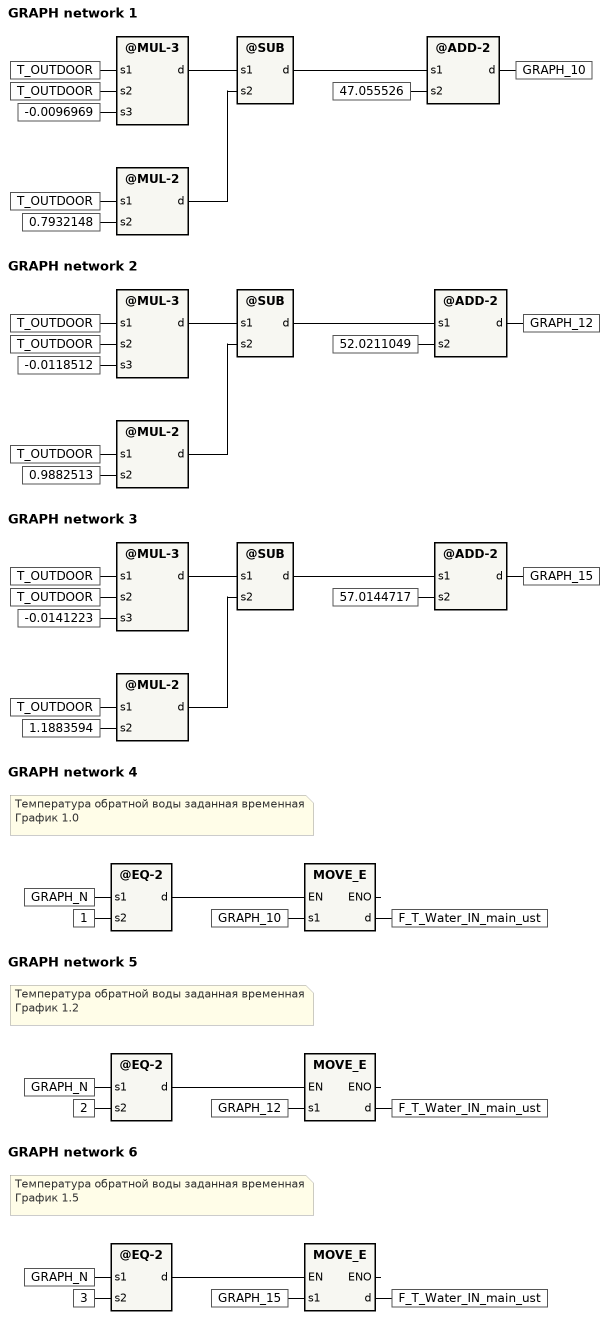
(* network 1 *)
GRAPH_10 := @ADD-2(@SUB(@MUL-3(T_OUTDOOR, T_OUTDOOR, -0.0096969), @MUL-2(T_OUTDOOR, 0.7932148)), 47.055526);
(* network 2 *)
GRAPH_12 := @ADD-2(@SUB(@MUL-3(T_OUTDOOR, T_OUTDOOR, -0.0118512), @MUL-2(T_OUTDOOR, 0.9882513)), 52.0211049);
(* network 3 *)
GRAPH_15 := @ADD-2(@SUB(@MUL-3(T_OUTDOOR, T_OUTDOOR, -0.0141223), @MUL-2(T_OUTDOOR, 1.1883594)), 57.0144717);
(* network 4 *)
(* Температура обратной воды заданная временная График 1.0 *)
MOVE_E(@EQ-2(GRAPH_N, 1), GRAPH_10, F_T_Water_IN_main_ust);
(* network 5 *)
(* Температура обратной воды заданная временная График 1.2 *)
MOVE_E(@EQ-2(GRAPH_N, 2), GRAPH_12, F_T_Water_IN_main_ust);
(* network 6 *)
(* Температура обратной воды заданная временная График 1.5 *)
MOVE_E(@EQ-2(GRAPH_N, 3), GRAPH_15, F_T_Water_IN_main_ust);
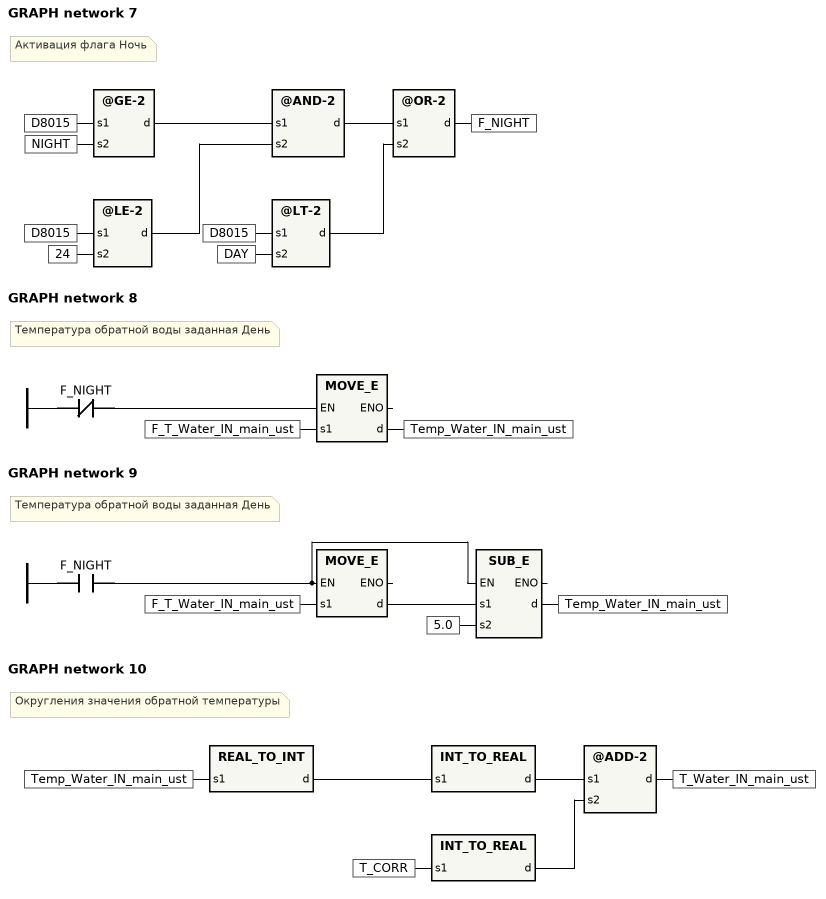
(* network 7 *)
(* Активация флага Ночь *)
F_NIGHT := @OR-2(@AND-2(@GE-2(D8015, NIGHT), @LE-2(D8015, 24)), @LT-2(D8015, DAY));
(* network 8 *)
(* Температура обратной воды заданная День *)
MOVE_E(NOT F_NIGHT, F_T_Water_IN_main_ust, Temp_Water_IN_main_ust);
(* network 9 *)
(* Температура обратной воды заданная День *)
MOVE_E(F_NIGHT, F_T_Water_IN_main_ust, _t1);
SUB_E(F_NIGHT, _t1, 5.0, Temp_Water_IN_main_ust);
(* network 10 *)
(* Округления значения обратной температуры *)
T_Water_IN_main_ust := @ADD-2(INT_TO_REAL(REAL_TO_INT(Temp_Water_IN_main_ust)), INT_TO_REAL(T_CORR));
END_FUNCTION_BLOCK

FUNCTION FUN_FILTER
VAR_INPUT
  InpF : REAL;
  OutF : REAL;
  Scan : INT;
  Tf : DINT;
END_VAR
VAR
  rScan : REAL;
  Param : REAL;
  FCorrect : BOOL;
  rTf : REAL;
  Output : REAL;
  TEMP1 : REAL;
  TEMP2 : REAL;
END_VAR
(* structured ladder/FBD written out as ST: instructions are called as NAME(EN, inputs, outputs); _pN, _eN, _tN stand for wires *)
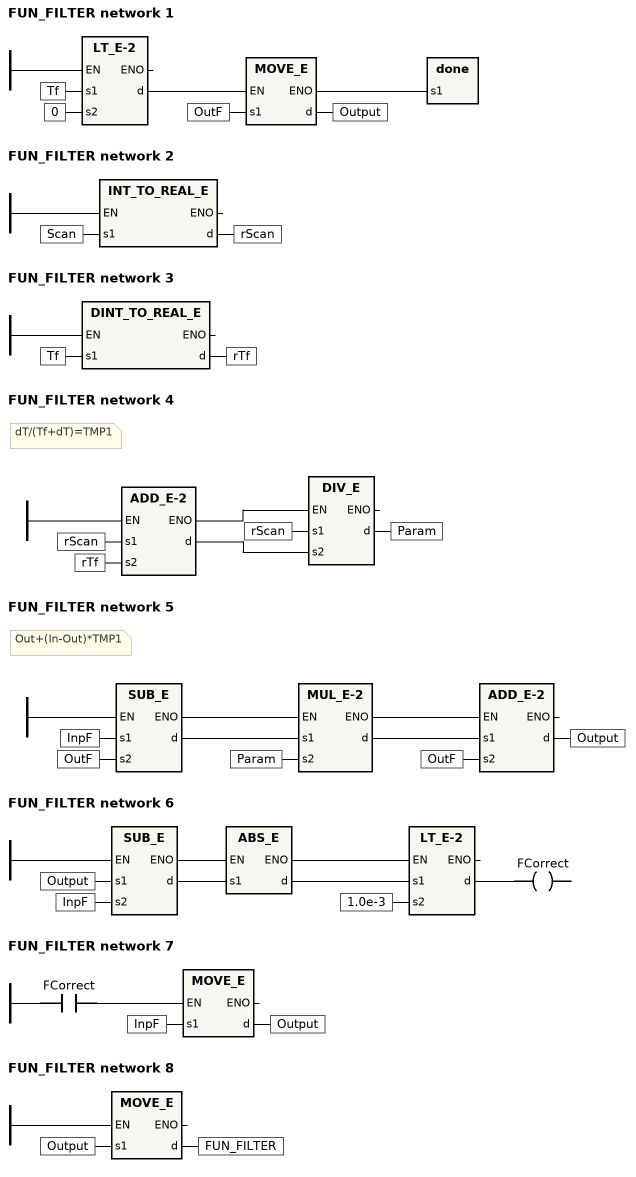
(* network 1 *)
LT_E(TRUE, Tf, 0, _t1);
_e2 := MOVE_E(_t1, OutF, Output);
(* element kind 9 done <- _e2 *)
(* network 2 *)
INT_TO_REAL_E(TRUE, Scan, rScan);
(* network 3 *)
DINT_TO_REAL_E(TRUE, Tf, rTf);
(* network 4 *)
(* dT/(Tf+dT)=TMP1 *)
_e2 := ADD_E(TRUE, rScan, rTf, _t1);
DIV_E(_e2, rScan, _t1, Param);
(* network 5 *)
(* Out+(In-Out)*TMP1 *)
_e2 := SUB_E(TRUE, InpF, OutF, _t1);
_e4 := MUL_E(_e2, _t1, Param, _t3);
ADD_E(_e4, _t3, OutF, Output);
(* network 6 *)
_e2 := SUB_E(TRUE, Output, InpF, _t1);
_e4 := ABS_E(_e2, _t1, _t3);
LT_E(_e4, _t3, 1.0e-3, _t5);
FCorrect := _t5;
(* network 7 *)
MOVE_E(FCorrect, InpF, Output);
(* network 8 done: *)
MOVE_E(TRUE, Output, FUN_FILTER);
END_FUNCTION

PROGRAM COUNTERS
VAR
  temp1 : BOOL;
  TON_1_1s : TON;
  time_sec : INT;
  time_min : INT;
  time_hour : INT;
  CIRC_PUMP_1_sec : INT;
  CIRC_PUMP_2_sec : INT;
  REZERV_PUMP_sec : INT;
  RECIRC_PUMP_12_sec : INT;
  TON_2_1s : TON;
  TON_3_1s : TON;
  TON_4_1s : TON;
  TON_5_1s : TON;
  BURNER_1_KOTEL_1_sec : INT;
  BURNER_2_KOTEL_1_sec : INT;
  BURNER_1_KOTEL_2_sec : INT;
  BURNER_2_KOTEL_2_sec : INT;
  TON_6_1s : TON;
  TON_7_1s : TON;
  TON_8_1s : TON;
END_VAR
(* structured ladder/FBD written out as ST: instructions are called as NAME(EN, inputs, outputs); _pN, _eN, _tN stand for wires *)
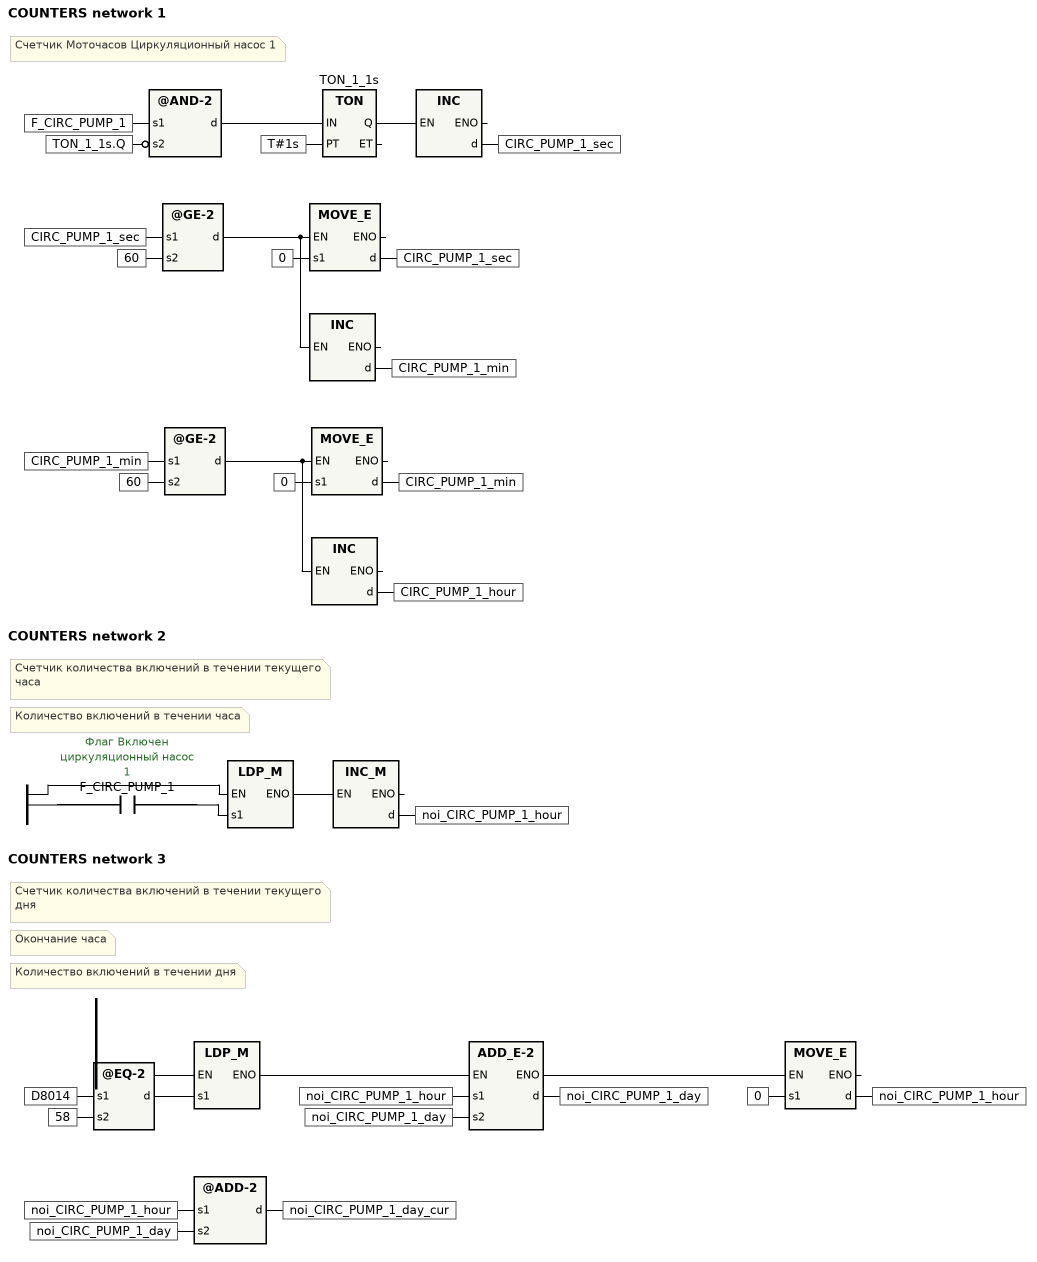
(* network 1 *)
(* Счетчик Моточасов Циркуляционный насос 1 *)
TON_1_1s(IN := @AND-2(F_CIRC_PUMP_1, NOT TON_1_1s.Q), PT := T#1s);
INC(TON_1_1s.Q, CIRC_PUMP_1_sec);
_p1 := @GE-2(CIRC_PUMP_1_sec, 60);
MOVE_E(_p1, 0, CIRC_PUMP_1_sec);
INC(_p1, CIRC_PUMP_1_min);
_p2 := @GE-2(CIRC_PUMP_1_min, 60);
MOVE_E(_p2, 0, CIRC_PUMP_1_min);
INC(_p2, CIRC_PUMP_1_hour);
(* network 2 *)
(* Счетчик количества включений в течении текущего часа *)
(* Количество включений в течении часа *)
_e1 := LDP_M(TRUE, F_CIRC_PUMP_1);
INC_M(_e1, noi_CIRC_PUMP_1_hour);
(* network 3 *)
(* Счетчик количества включений в течении текущего дня *)
(* Окончание часа *)
(* Количество включений в течении дня *)
_e1 := LDP_M(TRUE, @EQ-2(D8014, 58));
_e2 := ADD_E(_e1, noi_CIRC_PUMP_1_hour, noi_CIRC_PUMP_1_day, noi_CIRC_PUMP_1_day);
MOVE_E(_e2, 0, noi_CIRC_PUMP_1_hour);
noi_CIRC_PUMP_1_day_cur := @ADD-2(noi_CIRC_PUMP_1_hour, noi_CIRC_PUMP_1_day);
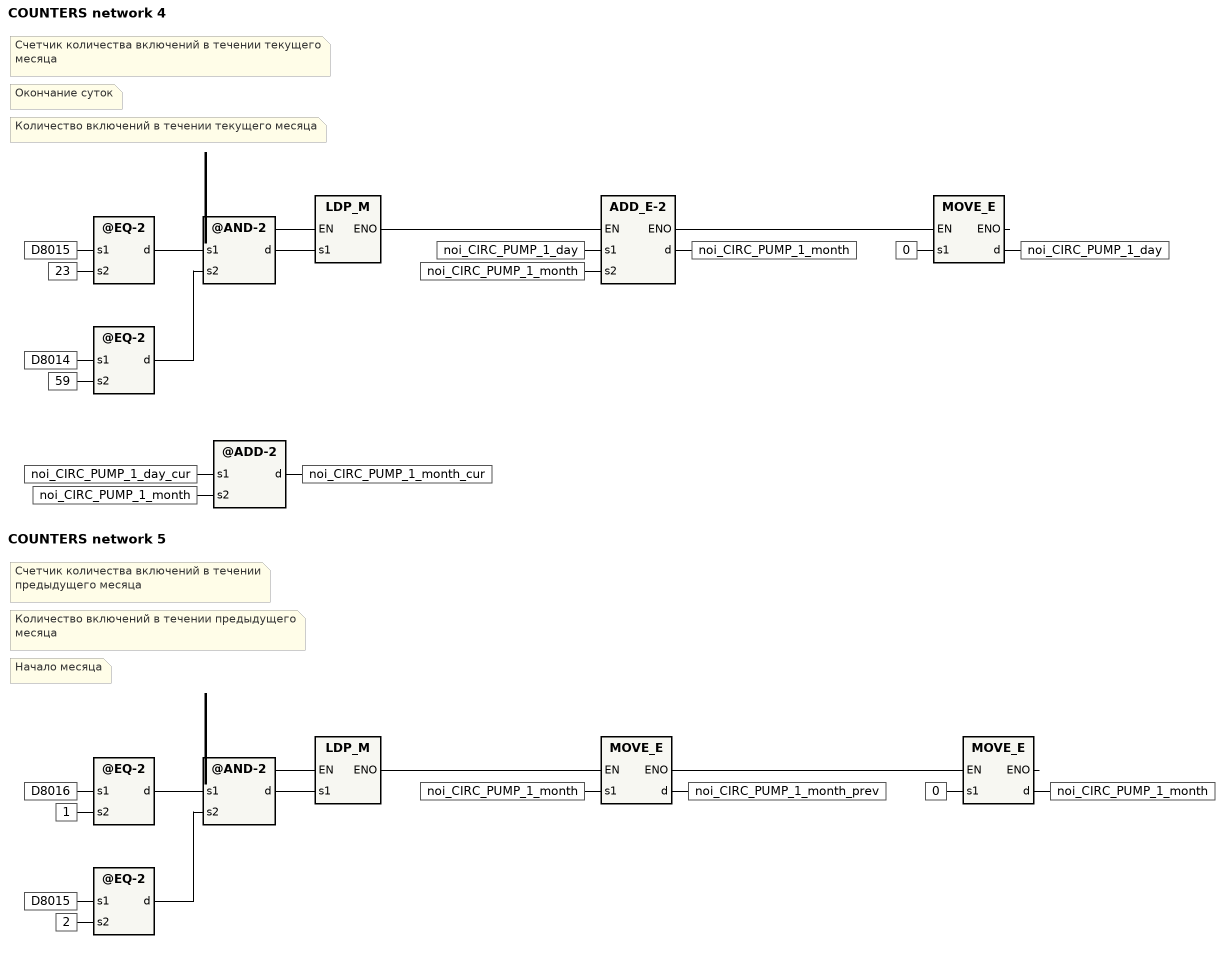
(* network 4 *)
(* Счетчик количества включений в течении текущего месяца *)
(* Окончание суток *)
(* Количество включений в течении текущего месяца *)
_e1 := LDP_M(TRUE, @AND-2(@EQ-2(D8015, 23), @EQ-2(D8014, 59)));
_e2 := ADD_E(_e1, noi_CIRC_PUMP_1_day, noi_CIRC_PUMP_1_month, noi_CIRC_PUMP_1_month);
MOVE_E(_e2, 0, noi_CIRC_PUMP_1_day);
noi_CIRC_PUMP_1_month_cur := @ADD-2(noi_CIRC_PUMP_1_day_cur, noi_CIRC_PUMP_1_month);
(* network 5 *)
(* Счетчик количества включений в течении предыдущего месяца *)
(* Количество включений в течении предыдущего месяца *)
(* Начало месяца *)
_e1 := LDP_M(TRUE, @AND-2(@EQ-2(D8016, 1), @EQ-2(D8015, 2)));
_e2 := MOVE_E(_e1, noi_CIRC_PUMP_1_month, noi_CIRC_PUMP_1_month_prev);
MOVE_E(_e2, 0, noi_CIRC_PUMP_1_month);
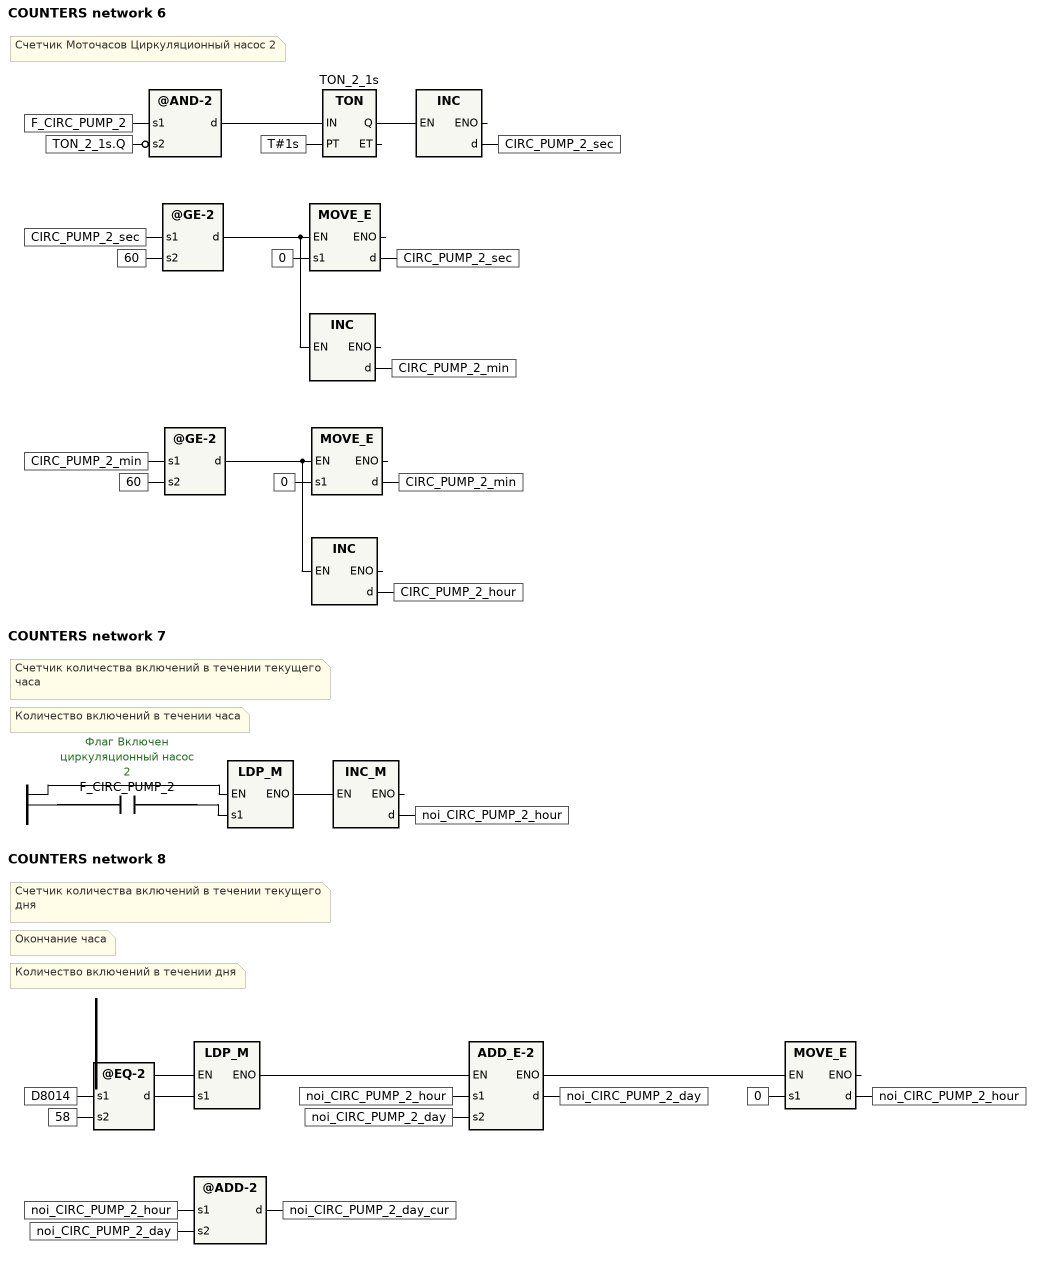
(* network 6 *)
(* Счетчик Моточасов Циркуляционный насос 2 *)
TON_2_1s(IN := @AND-2(F_CIRC_PUMP_2, NOT TON_2_1s.Q), PT := T#1s);
INC(TON_2_1s.Q, CIRC_PUMP_2_sec);
_p1 := @GE-2(CIRC_PUMP_2_sec, 60);
MOVE_E(_p1, 0, CIRC_PUMP_2_sec);
INC(_p1, CIRC_PUMP_2_min);
_p2 := @GE-2(CIRC_PUMP_2_min, 60);
MOVE_E(_p2, 0, CIRC_PUMP_2_min);
INC(_p2, CIRC_PUMP_2_hour);
(* network 7 *)
(* Счетчик количества включений в течении текущего часа *)
(* Количество включений в течении часа *)
_e1 := LDP_M(TRUE, F_CIRC_PUMP_2);
INC_M(_e1, noi_CIRC_PUMP_2_hour);
(* network 8 *)
(* Счетчик количества включений в течении текущего дня *)
(* Окончание часа *)
(* Количество включений в течении дня *)
_e1 := LDP_M(TRUE, @EQ-2(D8014, 58));
_e2 := ADD_E(_e1, noi_CIRC_PUMP_2_hour, noi_CIRC_PUMP_2_day, noi_CIRC_PUMP_2_day);
MOVE_E(_e2, 0, noi_CIRC_PUMP_2_hour);
noi_CIRC_PUMP_2_day_cur := @ADD-2(noi_CIRC_PUMP_2_hour, noi_CIRC_PUMP_2_day);
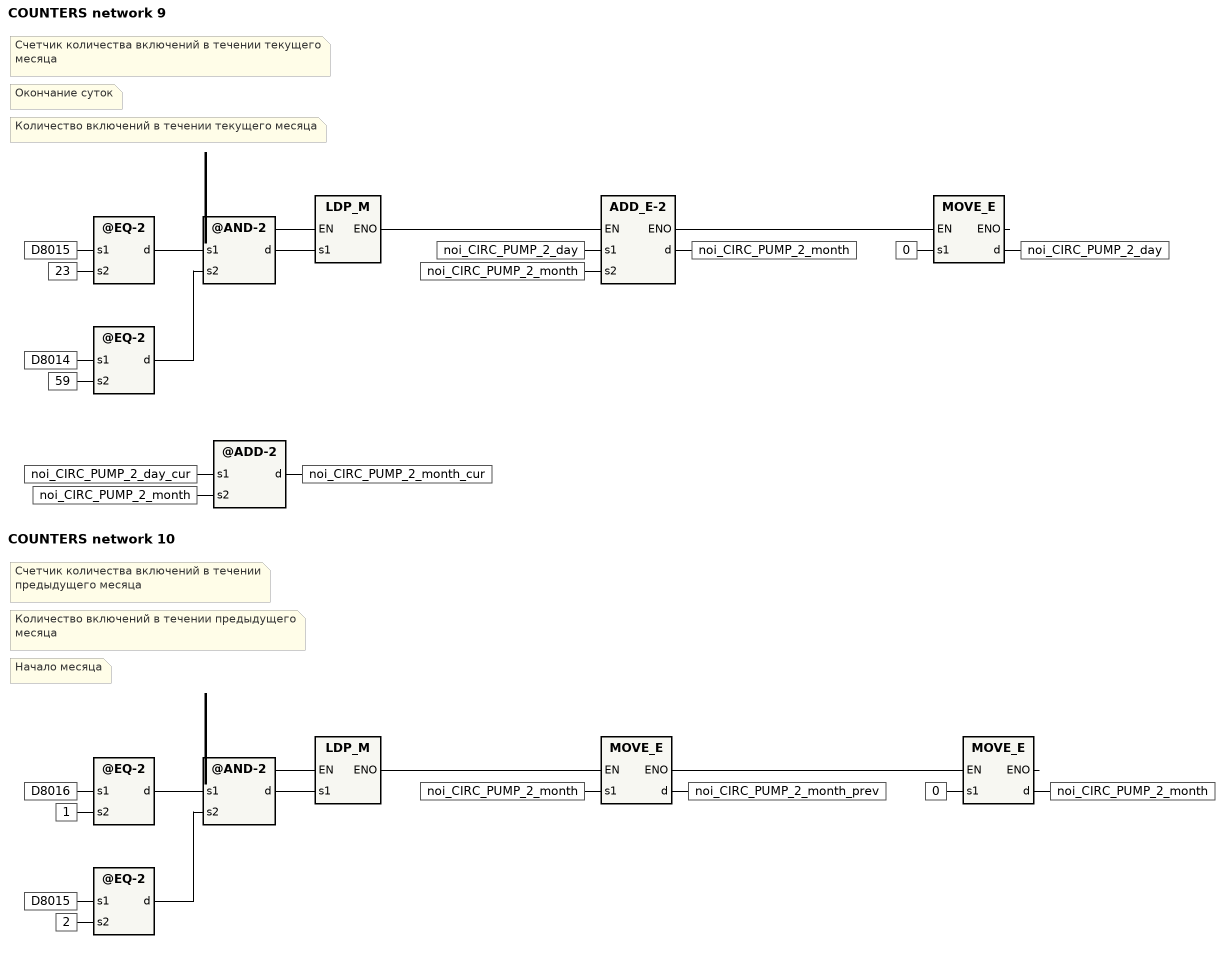
(* network 9 *)
(* Счетчик количества включений в течении текущего месяца *)
(* Окончание суток *)
(* Количество включений в течении текущего месяца *)
_e1 := LDP_M(TRUE, @AND-2(@EQ-2(D8015, 23), @EQ-2(D8014, 59)));
_e2 := ADD_E(_e1, noi_CIRC_PUMP_2_day, noi_CIRC_PUMP_2_month, noi_CIRC_PUMP_2_month);
MOVE_E(_e2, 0, noi_CIRC_PUMP_2_day);
noi_CIRC_PUMP_2_month_cur := @ADD-2(noi_CIRC_PUMP_2_day_cur, noi_CIRC_PUMP_2_month);
(* network 10 *)
(* Счетчик количества включений в течении предыдущего месяца *)
(* Количество включений в течении предыдущего месяца *)
(* Начало месяца *)
_e1 := LDP_M(TRUE, @AND-2(@EQ-2(D8016, 1), @EQ-2(D8015, 2)));
_e2 := MOVE_E(_e1, noi_CIRC_PUMP_2_month, noi_CIRC_PUMP_2_month_prev);
MOVE_E(_e2, 0, noi_CIRC_PUMP_2_month);
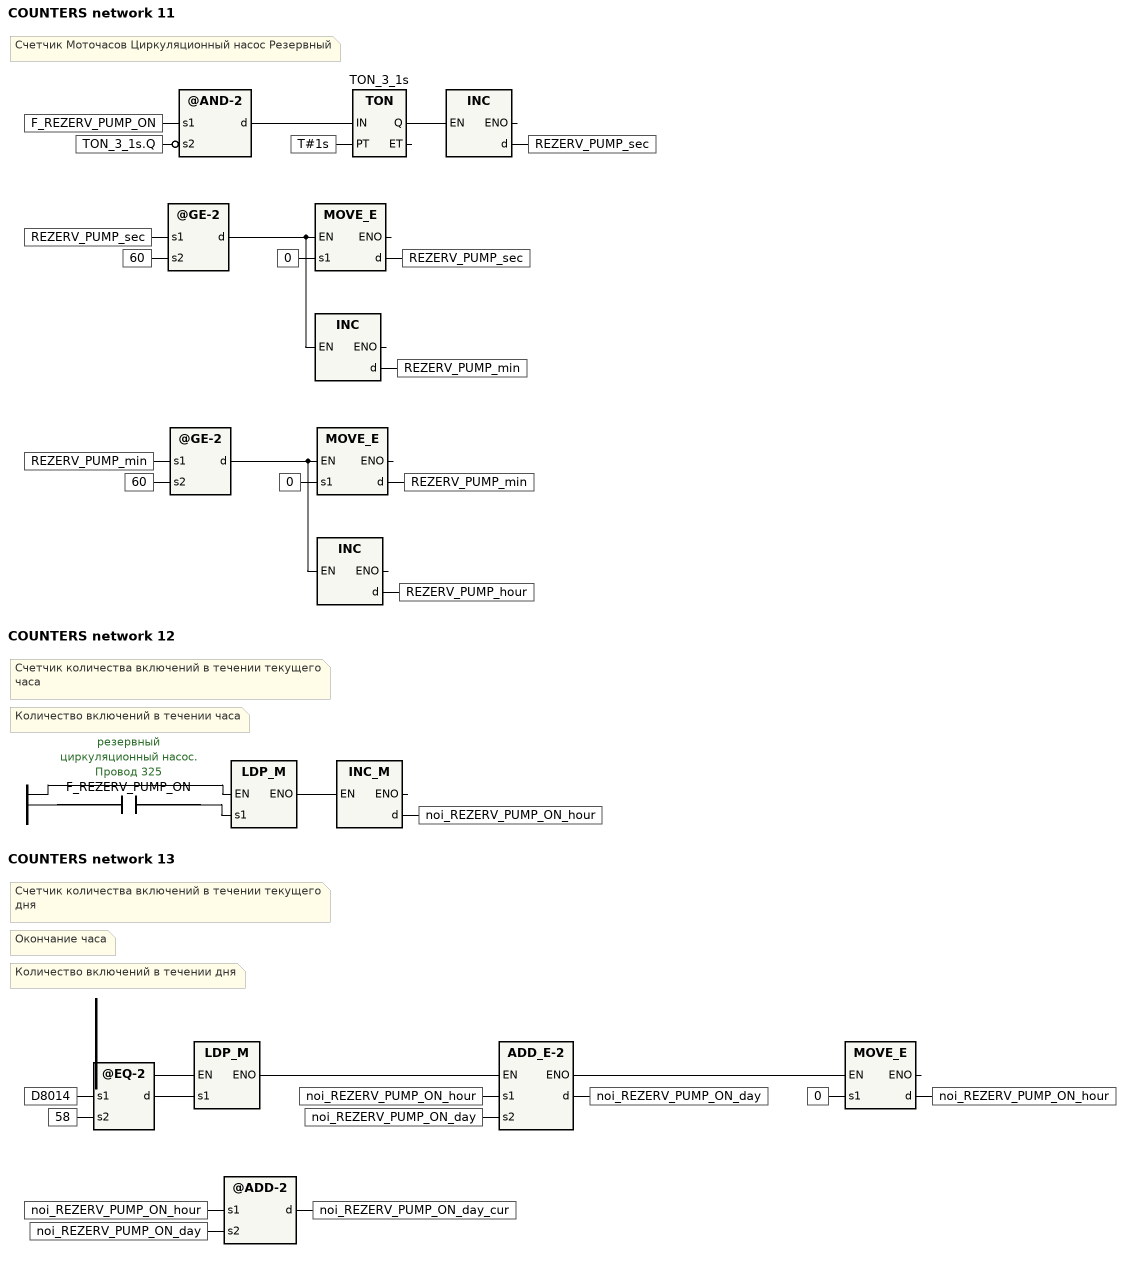
(* network 11 *)
(* Счетчик Моточасов Циркуляционный насос Резервный *)
TON_3_1s(IN := @AND-2(F_REZERV_PUMP_ON, NOT TON_3_1s.Q), PT := T#1s);
INC(TON_3_1s.Q, REZERV_PUMP_sec);
_p1 := @GE-2(REZERV_PUMP_sec, 60);
MOVE_E(_p1, 0, REZERV_PUMP_sec);
INC(_p1, REZERV_PUMP_min);
_p2 := @GE-2(REZERV_PUMP_min, 60);
MOVE_E(_p2, 0, REZERV_PUMP_min);
INC(_p2, REZERV_PUMP_hour);
(* network 12 *)
(* Счетчик количества включений в течении текущего часа *)
(* Количество включений в течении часа *)
_e1 := LDP_M(TRUE, F_REZERV_PUMP_ON);
INC_M(_e1, noi_REZERV_PUMP_ON_hour);
(* network 13 *)
(* Счетчик количества включений в течении текущего дня *)
(* Окончание часа *)
(* Количество включений в течении дня *)
_e1 := LDP_M(TRUE, @EQ-2(D8014, 58));
_e2 := ADD_E(_e1, noi_REZERV_PUMP_ON_hour, noi_REZERV_PUMP_ON_day, noi_REZERV_PUMP_ON_day);
MOVE_E(_e2, 0, noi_REZERV_PUMP_ON_hour);
noi_REZERV_PUMP_ON_day_cur := @ADD-2(noi_REZERV_PUMP_ON_hour, noi_REZERV_PUMP_ON_day);
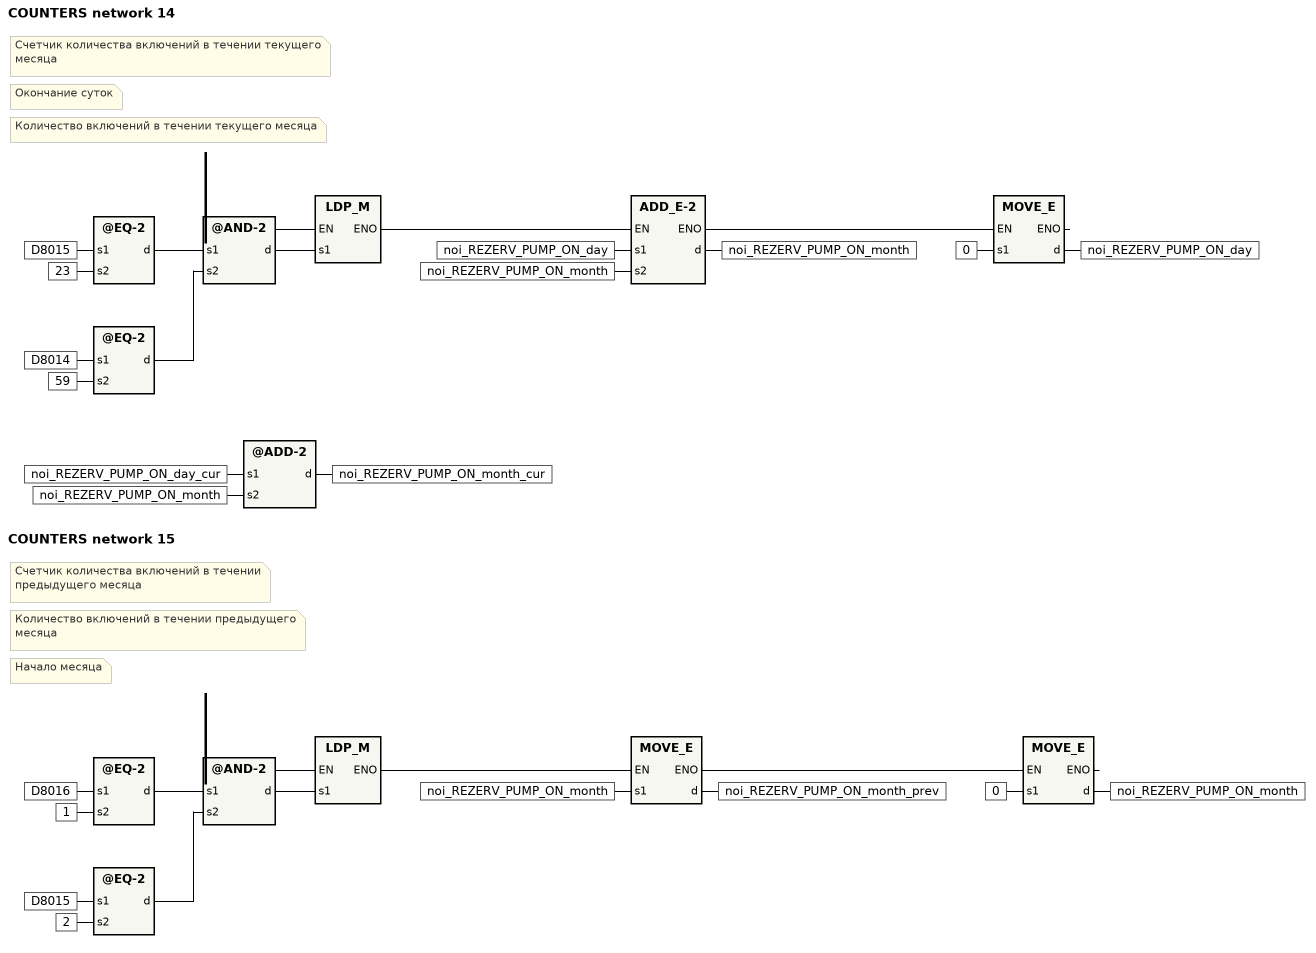
(* network 14 *)
(* Счетчик количества включений в течении текущего месяца *)
(* Окончание суток *)
(* Количество включений в течении текущего месяца *)
_e1 := LDP_M(TRUE, @AND-2(@EQ-2(D8015, 23), @EQ-2(D8014, 59)));
_e2 := ADD_E(_e1, noi_REZERV_PUMP_ON_day, noi_REZERV_PUMP_ON_month, noi_REZERV_PUMP_ON_month);
MOVE_E(_e2, 0, noi_REZERV_PUMP_ON_day);
noi_REZERV_PUMP_ON_month_cur := @ADD-2(noi_REZERV_PUMP_ON_day_cur, noi_REZERV_PUMP_ON_month);
(* network 15 *)
(* Счетчик количества включений в течении предыдущего месяца *)
(* Количество включений в течении предыдущего месяца *)
(* Начало месяца *)
_e1 := LDP_M(TRUE, @AND-2(@EQ-2(D8016, 1), @EQ-2(D8015, 2)));
_e2 := MOVE_E(_e1, noi_REZERV_PUMP_ON_month, noi_REZERV_PUMP_ON_month_prev);
MOVE_E(_e2, 0, noi_REZERV_PUMP_ON_month);
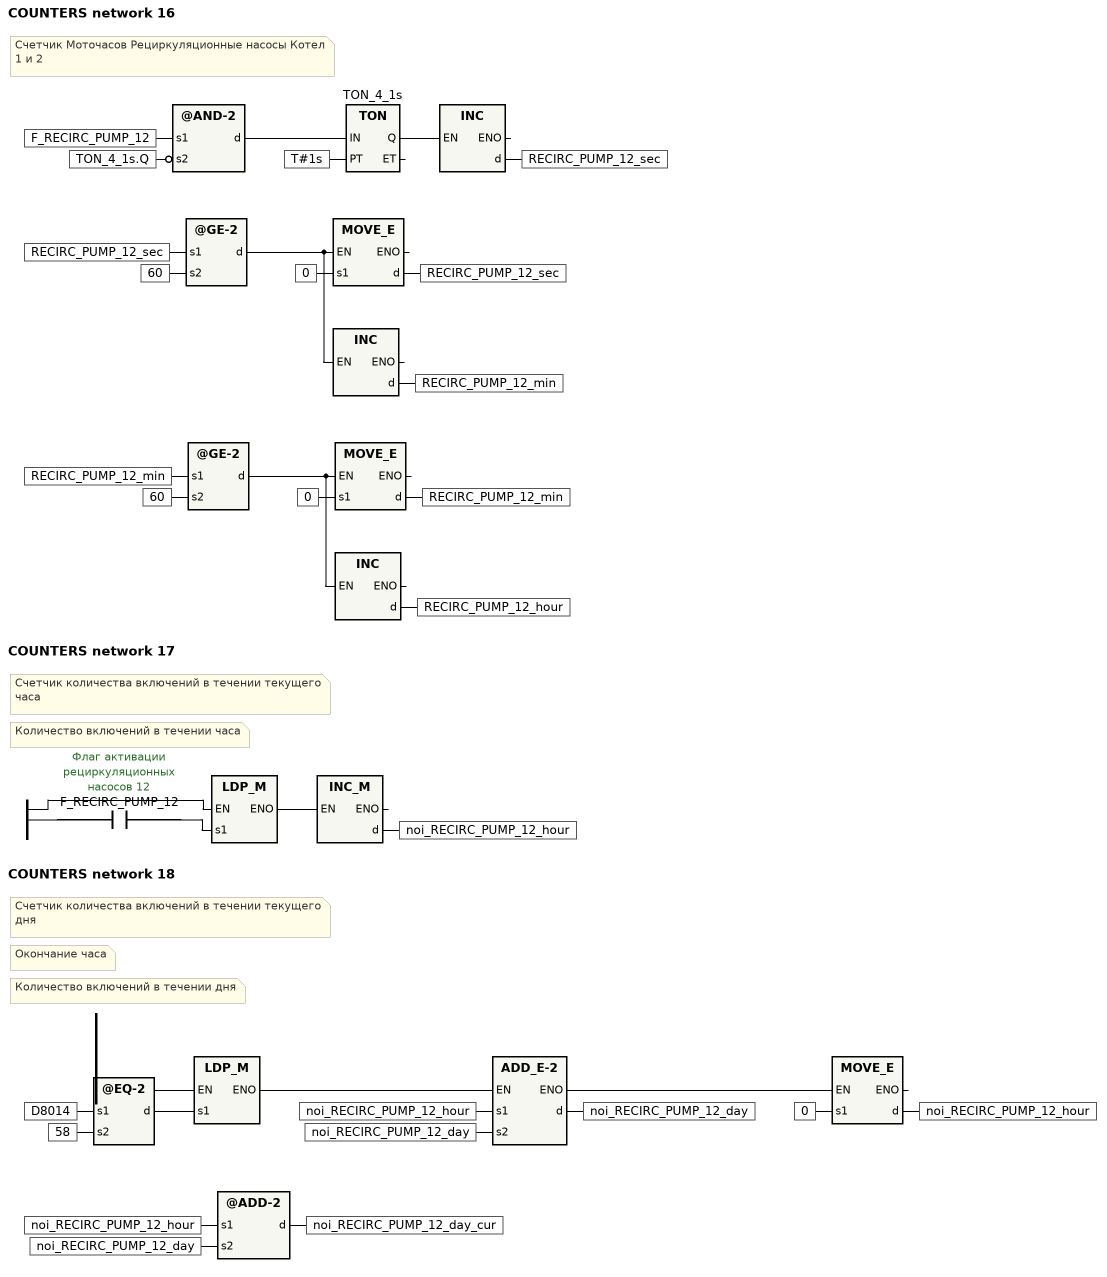
(* network 16 *)
(* Счетчик Моточасов Рециркуляционные насосы Котел 1 и 2 *)
TON_4_1s(IN := @AND-2(F_RECIRC_PUMP_12, NOT TON_4_1s.Q), PT := T#1s);
INC(TON_4_1s.Q, RECIRC_PUMP_12_sec);
_p1 := @GE-2(RECIRC_PUMP_12_sec, 60);
MOVE_E(_p1, 0, RECIRC_PUMP_12_sec);
INC(_p1, RECIRC_PUMP_12_min);
_p2 := @GE-2(RECIRC_PUMP_12_min, 60);
MOVE_E(_p2, 0, RECIRC_PUMP_12_min);
INC(_p2, RECIRC_PUMP_12_hour);
(* network 17 *)
(* Счетчик количества включений в течении текущего часа *)
(* Количество включений в течении часа *)
_e1 := LDP_M(TRUE, F_RECIRC_PUMP_12);
INC_M(_e1, noi_RECIRC_PUMP_12_hour);
(* network 18 *)
(* Счетчик количества включений в течении текущего дня *)
(* Окончание часа *)
(* Количество включений в течении дня *)
_e1 := LDP_M(TRUE, @EQ-2(D8014, 58));
_e2 := ADD_E(_e1, noi_RECIRC_PUMP_12_hour, noi_RECIRC_PUMP_12_day, noi_RECIRC_PUMP_12_day);
MOVE_E(_e2, 0, noi_RECIRC_PUMP_12_hour);
noi_RECIRC_PUMP_12_day_cur := @ADD-2(noi_RECIRC_PUMP_12_hour, noi_RECIRC_PUMP_12_day);
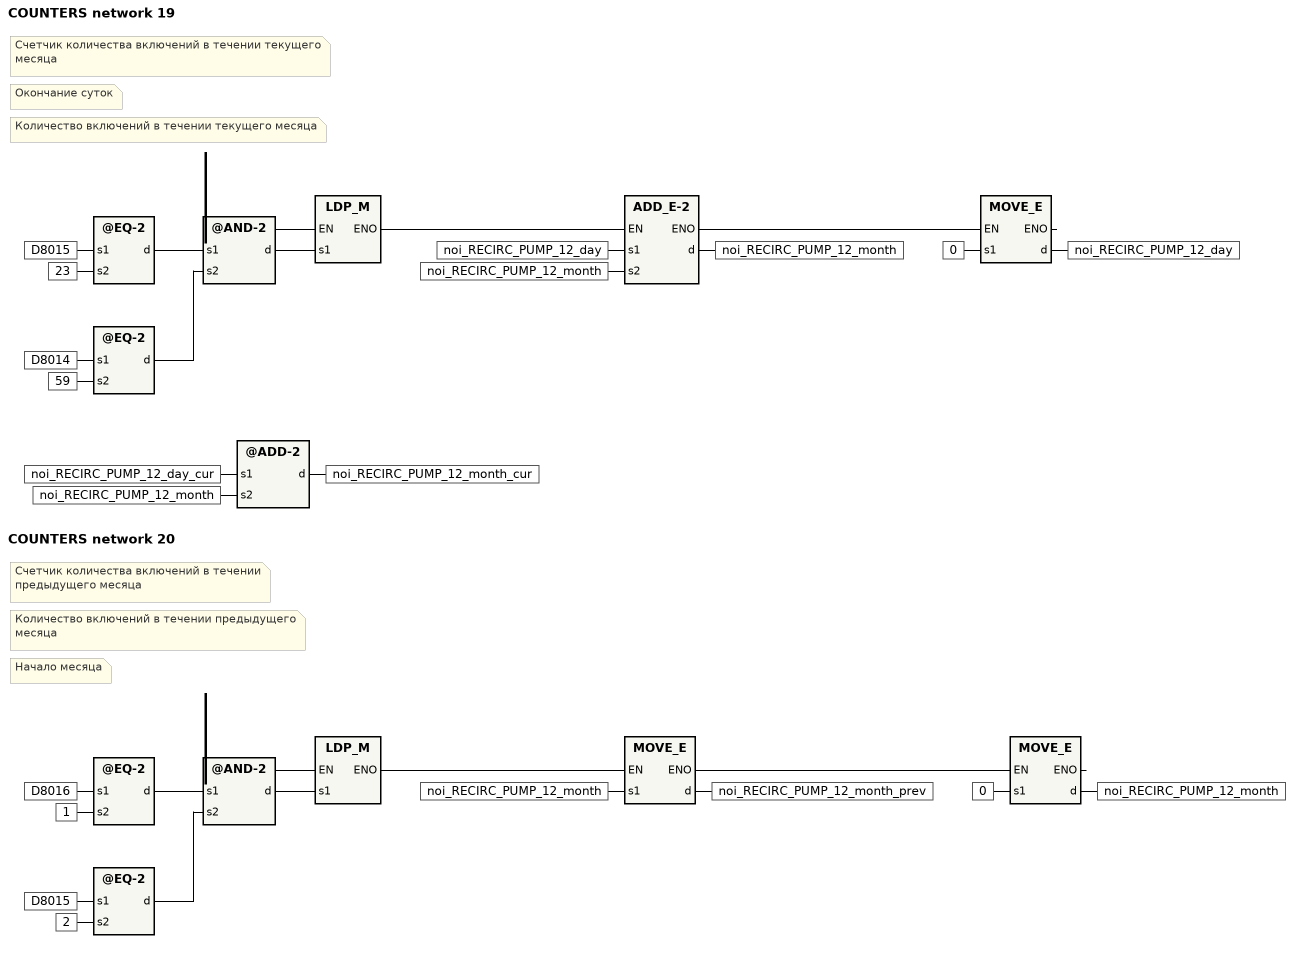
(* network 19 *)
(* Счетчик количества включений в течении текущего месяца *)
(* Окончание суток *)
(* Количество включений в течении текущего месяца *)
_e1 := LDP_M(TRUE, @AND-2(@EQ-2(D8015, 23), @EQ-2(D8014, 59)));
_e2 := ADD_E(_e1, noi_RECIRC_PUMP_12_day, noi_RECIRC_PUMP_12_month, noi_RECIRC_PUMP_12_month);
MOVE_E(_e2, 0, noi_RECIRC_PUMP_12_day);
noi_RECIRC_PUMP_12_month_cur := @ADD-2(noi_RECIRC_PUMP_12_day_cur, noi_RECIRC_PUMP_12_month);
(* network 20 *)
(* Счетчик количества включений в течении предыдущего месяца *)
(* Количество включений в течении предыдущего месяца *)
(* Начало месяца *)
_e1 := LDP_M(TRUE, @AND-2(@EQ-2(D8016, 1), @EQ-2(D8015, 2)));
_e2 := MOVE_E(_e1, noi_RECIRC_PUMP_12_month, noi_RECIRC_PUMP_12_month_prev);
MOVE_E(_e2, 0, noi_RECIRC_PUMP_12_month);
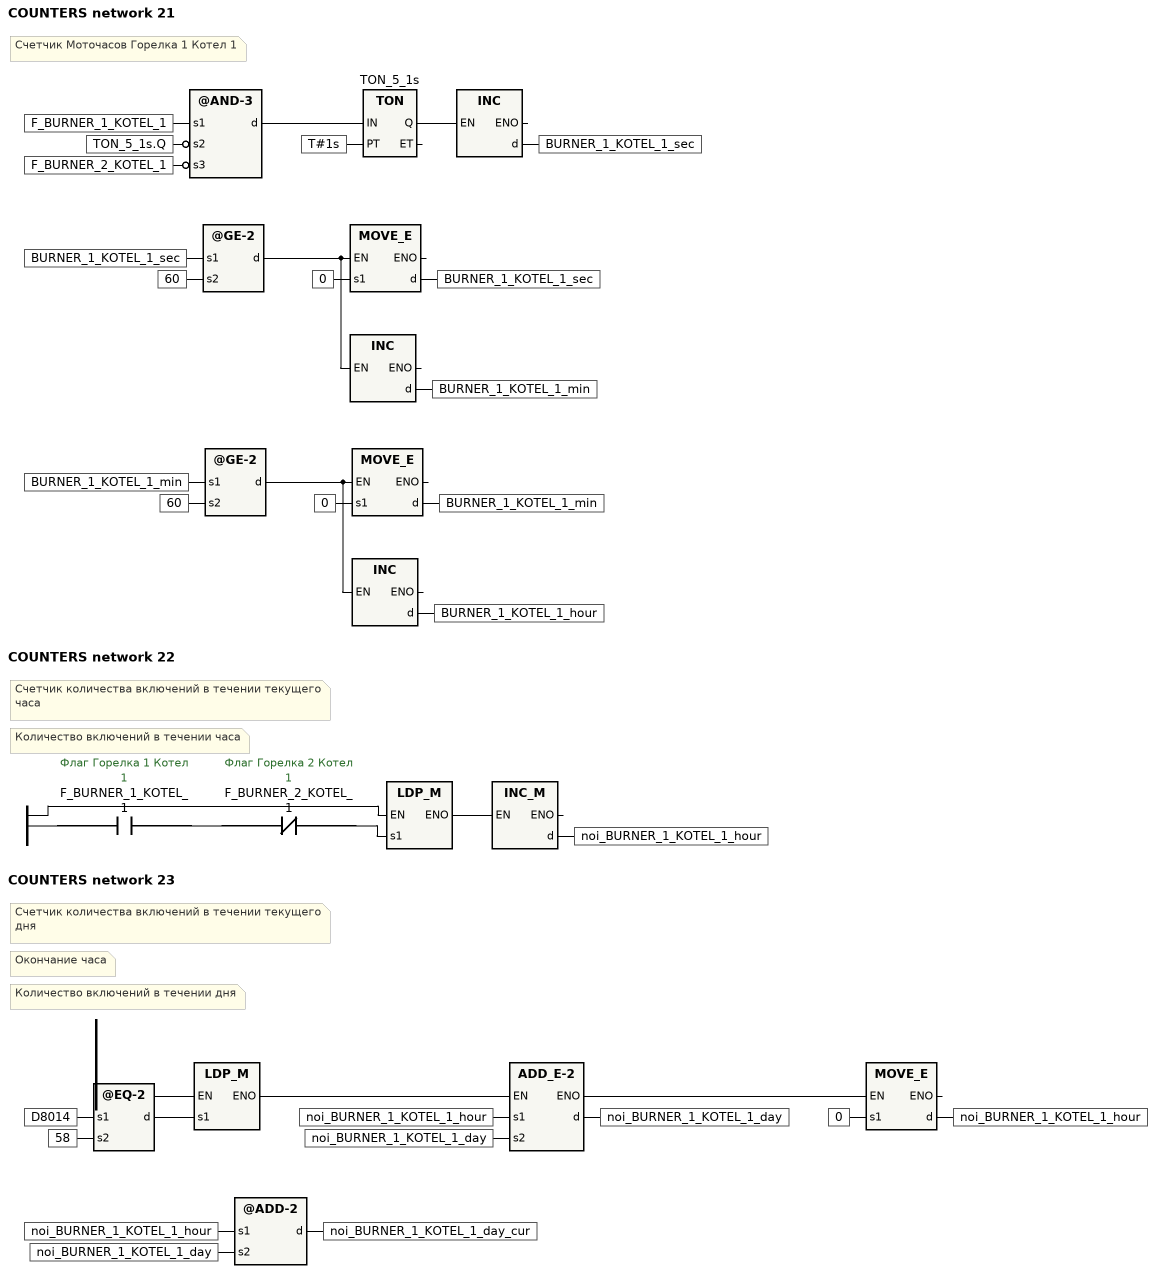
(* network 21 *)
(* Счетчик Моточасов Горелка 1 Котел 1 *)
TON_5_1s(IN := @AND-3(F_BURNER_1_KOTEL_1, NOT TON_5_1s.Q, NOT F_BURNER_2_KOTEL_1), PT := T#1s);
INC(TON_5_1s.Q, BURNER_1_KOTEL_1_sec);
_p1 := @GE-2(BURNER_1_KOTEL_1_sec, 60);
MOVE_E(_p1, 0, BURNER_1_KOTEL_1_sec);
INC(_p1, BURNER_1_KOTEL_1_min);
_p2 := @GE-2(BURNER_1_KOTEL_1_min, 60);
MOVE_E(_p2, 0, BURNER_1_KOTEL_1_min);
INC(_p2, BURNER_1_KOTEL_1_hour);
(* network 22 *)
(* Счетчик количества включений в течении текущего часа *)
(* Количество включений в течении часа *)
_e1 := LDP_M(TRUE, F_BURNER_1_KOTEL_1 AND NOT F_BURNER_2_KOTEL_1);
INC_M(_e1, noi_BURNER_1_KOTEL_1_hour);
(* network 23 *)
(* Счетчик количества включений в течении текущего дня *)
(* Окончание часа *)
(* Количество включений в течении дня *)
_e1 := LDP_M(TRUE, @EQ-2(D8014, 58));
_e2 := ADD_E(_e1, noi_BURNER_1_KOTEL_1_hour, noi_BURNER_1_KOTEL_1_day, noi_BURNER_1_KOTEL_1_day);
MOVE_E(_e2, 0, noi_BURNER_1_KOTEL_1_hour);
noi_BURNER_1_KOTEL_1_day_cur := @ADD-2(noi_BURNER_1_KOTEL_1_hour, noi_BURNER_1_KOTEL_1_day);
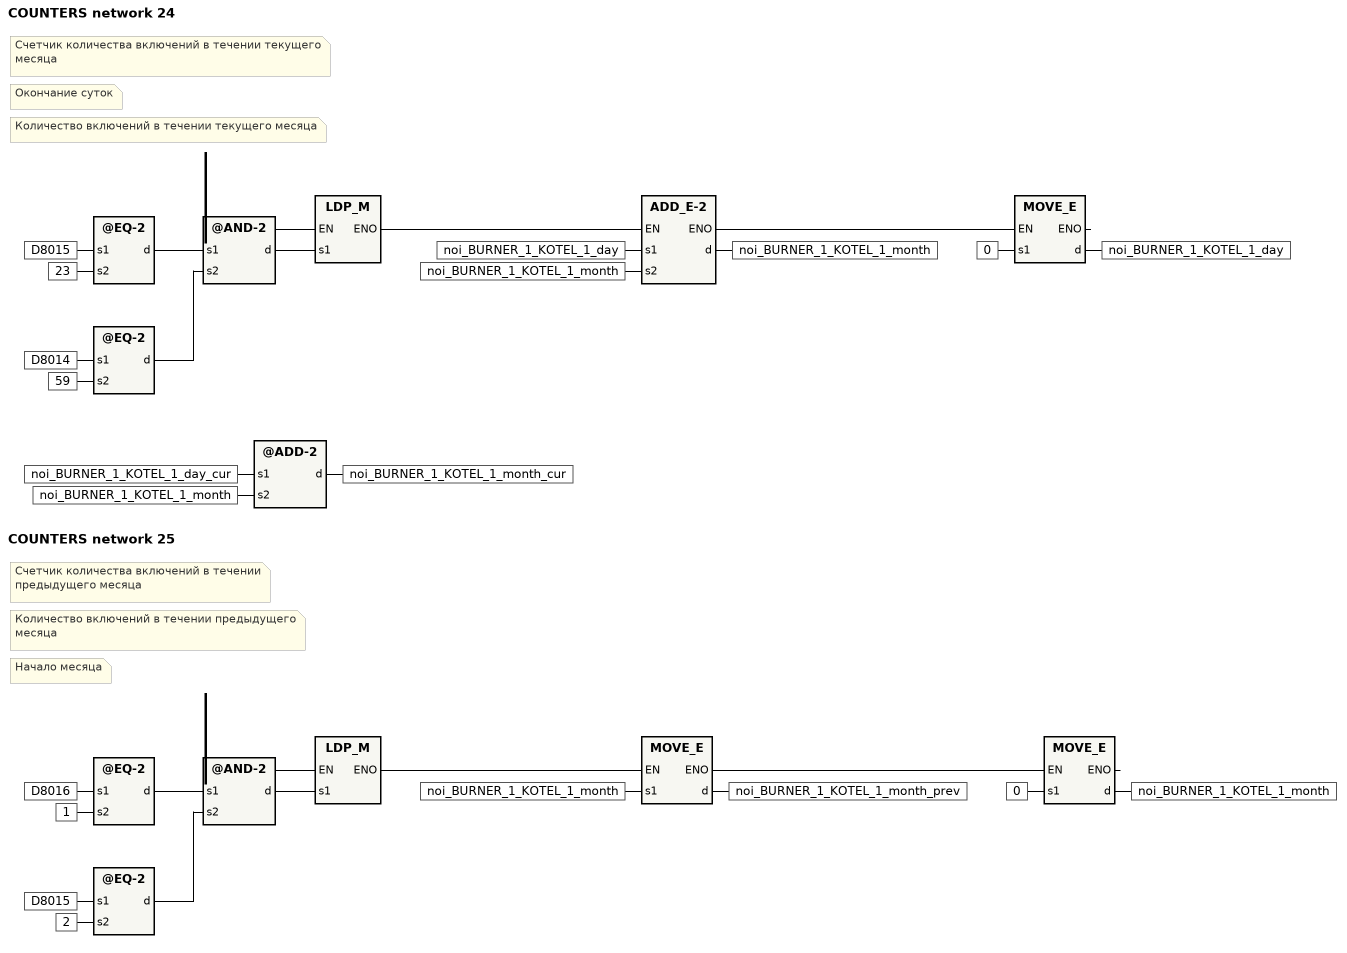
(* network 24 *)
(* Счетчик количества включений в течении текущего месяца *)
(* Окончание суток *)
(* Количество включений в течении текущего месяца *)
_e1 := LDP_M(TRUE, @AND-2(@EQ-2(D8015, 23), @EQ-2(D8014, 59)));
_e2 := ADD_E(_e1, noi_BURNER_1_KOTEL_1_day, noi_BURNER_1_KOTEL_1_month, noi_BURNER_1_KOTEL_1_month);
MOVE_E(_e2, 0, noi_BURNER_1_KOTEL_1_day);
noi_BURNER_1_KOTEL_1_month_cur := @ADD-2(noi_BURNER_1_KOTEL_1_day_cur, noi_BURNER_1_KOTEL_1_month);
(* network 25 *)
(* Счетчик количества включений в течении предыдущего месяца *)
(* Количество включений в течении предыдущего месяца *)
(* Начало месяца *)
_e1 := LDP_M(TRUE, @AND-2(@EQ-2(D8016, 1), @EQ-2(D8015, 2)));
_e2 := MOVE_E(_e1, noi_BURNER_1_KOTEL_1_month, noi_BURNER_1_KOTEL_1_month_prev);
MOVE_E(_e2, 0, noi_BURNER_1_KOTEL_1_month);